
           IF "Z256_Manager".tOutputData.rgxDataToProcessInter[#TMP_dIndexFAST] THEN

               #TMP_dEncoderOverFAST_cmm := #TMP_dEncValueFast - "Z256_Manager".tOutputData.rgdFireHeadThreshold_cmm[#TMP_dIndexFAST];

               //firing
               IF #TMP_dEncoderOverFAST_cmm >= 0 THEN



                   IF ("Z256_Manager".tOutputData.rgxFireHeadON_OFF[#TMP_dIndexFAST]) AND ("M256_Manag_IDB".M256F_IDB[#TMP_dIndexFAST].ST_xOutputEnable) AND
                       "M256_Manag_IDB".M256M_ST_xAllHeadPositioned AND "M256_Manag_IDB".M256A_IDB[#TMP_dIndexFAST].OUTPUT_xCarriageDescent THEN

                       "M256_Manag_IDB".M256F_IDB[#TMP_dIndexFAST].OUTPUT_xFireON := 1;

                   ELSE

                       "M256_Manag_IDB".M256F_IDB[#TMP_dIndexFAST].OUTPUT_xFireON := 0;

                   END_IF;

                   #TMP_xChangeFAST := 1;
                   "Z256_Manager".tOutputData.rgxDataToProcessInter[#TMP_dIndexFAST] := 0;
                   "M256_Manag_IDB".M256F_IDB[#TMP_dIndexFAST].AUX_dHeadMissionIDinProg := "Z256_Manager".tOutputData.dMissionCode;
                   "M256_Manag_IDB".M256F_IDB[#TMP_dIndexFAST].AUX_xHeadFiringMissionInProgress := "Z256_Manager".tOutputData.rgxFireHeadON_OFF[#TMP_dIndexFAST];

                   #TMP_xDummy := false;
                   FOR #TMP_dIndexFAST_2 := 0 TO "CONST_dNumberOfHeadsCycle" DO
                       IF "Z256_Manager".tOutputData.rgxFireHeadON_OFF[#TMP_dIndexFAST_2] THEN
                           #TMP_xDummy := true;
                       END_IF;
                   END_FOR;
                   IF NOT (#TMP_xDummy) THEN
                       "M256_Manag_IDB".M256F_IDB[#TMP_dIndexFAST].AUX_dHeadMissionIDinProg := 0;
                   END_IF;
               END_IF;
           END_IF;
       END_FOR;


       #TMP_xDummy := false;
       FOR #TMP_dIndexFAST := 0 TO "CONST_dNumberOfHeadsCycle" DO
           IF "Z256_Manager".tOutputData.rgxDataToProcessInter[#TMP_dIndexFAST] <> 0 THEN
               #TMP_xDummy := true;
           END_IF;
       END_FOR;
       IF #TMP_xDummy = false THEN
           "Z256_Manager".tOutputData.xGateOpen := 0;
       END_IF;
       //Immagine di processo aggiornata automaticamente con l'OB
       //    IF #TMP_xChangeFAST THEN
       //        #TMP_iRetVal:=UPDAT_PO(PART := "IPP 1", FLADDR => "DEBUG_FiringAdressError");
       //    END_IF;


   END_IF;


   "o.1B160AP1.EnableCard1":=  "M256_Manag_IDB".M256F_IDB[0].OUTPUT_xFireON OR"M256_Manag_IDB".M256F_IDB[0].INPUT_xForceFiring;
   "o.1B160AP1.EnableCard2" := "M256_Manag_IDB".M256F_IDB[1].OUTPUT_xFireON OR "M256_Manag_IDB".M256F_IDB[1].INPUT_xForceFiring;
   "o.1B160AP1.EnableCard3" := "M256_Manag_IDB".M256F_IDB[2].OUTPUT_xFireON OR "M256_Manag_IDB".M256F_IDB[2].INPUT_xForceFiring;
   "o.1B160AP1.EnableCard4" := "M256_Manag_IDB".M256F_IDB[3].OUTPUT_xFireON OR "M256_Manag_IDB".M256F_IDB[3].INPUT_xForceFiring;
   "o.1B160AP1.EnableCard5" := "M256_Manag_IDB".M256F_IDB[4].OUTPUT_xFireON OR "M256_Manag_IDB".M256F_IDB[4].INPUT_xForceFiring;
   "o.1B160AP1.EnableCard5" := "M256_Manag_IDB".M256F_IDB[5].OUTPUT_xFireON OR "M256_Manag_IDB".M256F_IDB[4].INPUT_xForceFiring;
   "o.1B160AP1.EnableCard5" := "M256_Manag_IDB".M256F_IDB[6].OUTPUT_xFireON OR "M256_Manag_IDB".M256F_IDB[4].INPUT_xForceFiring;
   "o.1B160AP1.EnableCard5" := "M256_Manag_IDB".M256F_IDB[7].OUTPUT_xFireON OR "M256_Manag_IDB".M256F_IDB[4].INPUT_xForceFiring;
END_REGION
END_ORGANIZATION_BLOCK

ORGANIZATION_BLOCK "Startup"   // OB100, SCL, Startup
TITLE = "Complete Restart"
{ S7_Optimized_Access := 'TRUE' }
VERSION : 0.1
   VAR_INPUT
      LostRetentive : Bool;   // True if retentive data are lost
      LostRTC : Bool;   // True if date and time are lost
   END_VAR
   VAR_TEMP
      TMP_dIndex : DInt;
   END_VAR
BEGIN
   // Start Auto Sequence after PLC restart

   "OB_Initialize".IN_xInitialize := TRUE;

   "INIT_PlantCostants"();

   //FORCE MANUAL STATE
   "Z256_hmi".tHMW.xGeneralReset := 1;

   FOR #TMP_dIndex := 0 TO "CONST_dNumberOfHeadsCycle" DO
       "M256_Manag_IDB".M256M_IDB[#TMP_dIndex].ST_xHeadInitialized := 0;
       "M256_Manag_IDB".M256M_IDB[#TMP_dIndex].AUX_dHeadRequestPosition_cmm := "M256_Manag_IDB".M256M_IDB[#TMP_dIndex].tHMR.dHeadHomePositions_cmm; 
       "Z256_hmi".tHMW.rgxHeadEnabled[#TMP_dIndex] := true;
   END_FOR;
END_ORGANIZATION_BLOCK

// folder: 07_ArrayScada

FUNCTION "SCADA_Mapping" : Void   // FC8, SCL
{ S7_Optimized_Access := 'TRUE' }
VERSION : 0.1
   VAR_TEMP
      TMP_dIndex : DInt;
   END_VAR
BEGIN

   //Move Z256 HMR
   "DB_Z256_Scada".tHMR.xCalibrationsAllowed:="Z256_hmi".tHMR.xCalibrationsAllowed;
   "DB_Z256_Scada".tHMR.xZoneAlarm:="Z256_hmi".tHMR.xZoneAlarm;
   "DB_Z256_Scada".tHMR.dZoneMode:="Z256_hmi".tHMR.dZoneMode;

   "DB_Z256_Scada".tHMR.dCabinetStatusMCC:="Z256_hmi".tHMR.dCabinetStatus;
   "DB_Z256_Scada".tHMR.dProdModeRequest:="Z256_hmi".tHMR.dProdModeRequest;
   "DB_Z256_Scada".tHMR.dProdModeActual:="Z256_hmi".tHMR.dProdModeActual;

   "DB_Z256_Scada".tHMR."rgdHeadsActualStatus[0]":="Z256_hmi".tHMR.rgdHeadsActualStatus[0];
   "DB_Z256_Scada".tHMR."rgdHeadsActualStatus[1]":="Z256_hmi".tHMR.rgdHeadsActualStatus[1];
   "DB_Z256_Scada".tHMR."rgdHeadsActualStatus[2]":="Z256_hmi".tHMR.rgdHeadsActualStatus[2];
   "DB_Z256_Scada".tHMR."rgdHeadsActualStatus[3]":="Z256_hmi".tHMR.rgdHeadsActualStatus[3];
   "DB_Z256_Scada".tHMR."rgdHeadsActualStatus[4]":="Z256_hmi".tHMR.rgdHeadsActualStatus[4];
   "DB_Z256_Scada".tHMR."rgdHeadsActualStatus[5]":="Z256_hmi".tHMR.rgdHeadsActualStatus[5];
   "DB_Z256_Scada".tHMR."rgdHeadsActualStatus[6]":="Z256_hmi".tHMR.rgdHeadsActualStatus[6];
   "DB_Z256_Scada".tHMR."rgdHeadsActualStatus[7]":="Z256_hmi".tHMR.rgdHeadsActualStatus[7];


   //Move Z256 HMW
   //
   "Z256_hmi".tHMW.xFaultsReset:="DB_Z256_Scada".tHMW.xFaultsReset ;
   "Z256_hmi".tHMW.xAutoModeReq:= "DB_Z256_Scada".tHMW.xAutoModeReq ;
   "Z256_hmi".tHMW.xGeneralReset:= "DB_Z256_Scada".tHMW.xGeneralReset ;
   "Z256_hmi".tHMW.xCutOnBreakEnabled:="DB_Z256_Scada".tHMW.xCutOnBreakEnabled  ;
   "Z256_hmi".tHMW.xManModeReq := "DB_Z256_Scada".tHMW.xManModeReq;
   "Z256_hmi".tHMW.xMotorsAndCardsInitialize:= "DB_Z256_Scada".tHMW.xMotorsAndCardsInitialize ;
   "Z256_hmi".tHMW.xOutOfProdReq:= "DB_Z256_Scada".tHMW.xOutOfProdReq ;
   "Z256_hmi".tHMW.xInProdReq:= "DB_Z256_Scada".tHMW.xInProdReq   ;
   "Z256_hmi".tHMW.xPositionCalibrationRequest := "DB_Z256_Scada".tHMW.xPositionCalibrationRequest;
   "Z256_hmi".tHMW.xForceHeadsHoming:= "DB_Z256_Scada".tHMW.xForceHeadsHoming   ;
   "Z256_hmi".tHMW.xBridgeOffsetCalibrationRequest:="DB_Z256_Scada".tHMW.xBridgeOffsetCalibrationRequest;
   "Z256_hmi".tHMW.tManCmd.xBrakeEngage:="DB_Z256_Scada".tHMW.tManCmd.xBrakeEngage;
   "Z256_hmi".tHMW.tManCmd.xBrakeRelease:="DB_Z256_Scada".tHMW.tManCmd.xBrakeRelease;

   "Z256_hmi".tHMW.rgxHeadEnabled[0] := "DB_Z256_Scada".tHMW.xHeadEnabled_1;
   "Z256_hmi".tHMW.rgxHeadEnabled[1] := "DB_Z256_Scada".tHMW.xHeadEnabled_2;
   "Z256_hmi".tHMW.rgxHeadEnabled[2] := "DB_Z256_Scada".tHMW.xHeadEnabled_3;
   "Z256_hmi".tHMW.rgxHeadEnabled[3] := "DB_Z256_Scada".tHMW.xHeadEnabled_4;
   "Z256_hmi".tHMW.rgxHeadEnabled[4] := "DB_Z256_Scada".tHMW.xHeadEnabled_5;
   "Z256_hmi".tHMW.rgxHeadEnabled[5] := "DB_Z256_Scada".tHMW.xHeadEnabled_6;
   "Z256_hmi".tHMW.rgxHeadEnabled[6] := "DB_Z256_Scada".tHMW.xHeadEnabled_7;
   "Z256_hmi".tHMW.rgxHeadEnabled[7] := "DB_Z256_Scada".tHMW.xHeadEnabled_8;

   "Z256_hmi".tHMW.dMoveBridgeOffset_cmm := "DB_Z256_Scada".tHMW.dMoveBridgeOffset_cmm;
   "Z256_hmi".tHMW.dNumberOfLites := "DB_Z256_Scada".tHMW.dNumberOfLites;
   "Z256_hmi".tHMW.dPressureScalerOnSample_perc := "DB_Z256_Scada".tHMW.dPressureScalerOnSample_perc;

   "Z256_hmi".tHMW.rgdHeadSelected[0]:="DB_Z256_Scada".tHMW.dHead_Selected_1;
   "Z256_hmi".tHMW.rgdHeadSelected[1]:="DB_Z256_Scada".tHMW.dHead_Selected_2;
   "Z256_hmi".tHMW.rgdHeadSelected[2]:="DB_Z256_Scada".tHMW.dHead_Selected_3;
   "Z256_hmi".tHMW.rgdHeadSelected[3]:="DB_Z256_Scada".tHMW.dHead_Selected_4;
   "Z256_hmi".tHMW.rgdHeadSelected[4]:="DB_Z256_Scada".tHMW.dHead_Selected_5;
   "Z256_hmi".tHMW.rgdHeadSelected[5]:="DB_Z256_Scada".tHMW.dHead_Selected_6;
   "Z256_hmi".tHMW.rgdHeadSelected[6]:="DB_Z256_Scada".tHMW.dHead_Selected_7;
   "Z256_hmi".tHMW.rgdHeadSelected[7] :="DB_Z256_Scada".tHMW.dHead_Selected_8;

   "Z256_hmi".tHMW.rgdCutWidthTeo_cmm[0] := "DB_Z256_Scada".tHMW.dCutWidthTeo_cmm_1;
   "Z256_hmi".tHMW.rgdCutWidthTeo_cmm[1] := "DB_Z256_Scada".tHMW.dCutWidthTeo_cmm_2;
   "Z256_hmi".tHMW.rgdCutWidthTeo_cmm[2] := "DB_Z256_Scada".tHMW.dCutWidthTeo_cmm_3;
   "Z256_hmi".tHMW.rgdCutWidthTeo_cmm[3] := "DB_Z256_Scada".tHMW."dCutWidthTeo_cmm_4";
   "Z256_hmi".tHMW.rgdCutWidthTeo_cmm[4] := "DB_Z256_Scada".tHMW."dCutWidthTeo_cmm_5";
   "Z256_hmi".tHMW.rgdCutWidthTeo_cmm[5] := "DB_Z256_Scada".tHMW."dCutWidthTeo_cmm_6";
   "Z256_hmi".tHMW.rgdCutWidthTeo_cmm[6] := "DB_Z256_Scada".tHMW."dCutWidthTeo_cmm_7";
   "Z256_hmi".tHMW.rgdCutWidthTeo_cmm[7] := "DB_Z256_Scada".tHMW."dCutWidthTeo_cmm_8";


   "Z256_hmi".tHMW.rgdCutWidthReal_cmm[0]:="DB_Z256_Scada".tHMW.dCutWidthReal_cmm_1;
   "Z256_hmi".tHMW.rgdCutWidthReal_cmm[1]:="DB_Z256_Scada".tHMW.dCutWidthReal_cmm_2;
   "Z256_hmi".tHMW.rgdCutWidthReal_cmm[2]:="DB_Z256_Scada".tHMW.dCutWidthReal_cmm_3;
   "Z256_hmi".tHMW.rgdCutWidthReal_cmm[3]:="DB_Z256_Scada".tHMW."dCutWidthReal_cmm_4";
   "Z256_hmi".tHMW.rgdCutWidthReal_cmm[4]:="DB_Z256_Scada".tHMW."dCutWidthReal_cmm_5";
   "Z256_hmi".tHMW.rgdCutWidthReal_cmm[5]:="DB_Z256_Scada".tHMW."dCutWidthReal_cmm_6";
   "Z256_hmi".tHMW.rgdCutWidthReal_cmm[6]:="DB_Z256_Scada".tHMW."dCutWidthReal_cmm_7";
   "Z256_hmi".tHMW.rgdCutWidthReal_cmm[7]:="DB_Z256_Scada".tHMW."dCutWidthTeo_cmm_8";

   (* //Move Z256 ALM
   "DB_M256M_Scada".tAlm.tS.tS0 := "DB_Z256_Scada".tAlm.tS.tS0;
   "DB_Z256_Scada".tAlm.tS.tS0.x0 := "DB_Z256_Scada".tAlm.tS.tS0.x0;
   "DB_Z256_Scada".tAlm.tS.tS0.x1 := "DB_Z256_Scada".tAlm.tS.tS0.x1;
   "DB_Z256_Scada".tAlm.tS.tS0.x2 := "DB_Z256_Scada".tAlm.tS.tS0.x2;
   "DB_Z256_Scada".tAlm.tS.tS0.x3 := "DB_Z256_Scada".tAlm.tS.tS0.x3;
   "DB_Z256_Scada".tAlm.tS.tS0.x4 := "DB_Z256_Scada".tAlm.tS.tS0.x4;
   "DB_Z256_Scada".tAlm.tS.tS0.x5 := "DB_Z256_Scada".tAlm.tS.tS0.x5;
   "DB_Z256_Scada".tAlm.tS.tS0.x6 := "DB_Z256_Scada".tAlm.tS.tS0.x6;
   "DB_Z256_Scada".tAlm.tS.tS0.x7 := "DB_Z256_Scada".tAlm.tS.tS0.x7;
   "DB_Z256_Scada".tAlm.tS.tS0.x8 := "DB_Z256_Scada".tAlm.tS.tS0.x8;

   "DB_Z256_Scada".tAlm.tS.tS0.x9 := "DB_Z256_Scada".tAlm.tS.tS0.x9;
   "DB_Z256_Scada".tAlm.tS.tS0.x10 := "DB_Z256_Scada".tAlm.tS.tS0.x10;
   "DB_Z256_Scada".tAlm.tS.tS0.x11 := "DB_Z256_Scada".tAlm.tS.tS0.x11;
   "DB_Z256_Scada".tAlm.tS.tS0.x12 := "DB_Z256_Scada".tAlm.tS.tS0.x12;
   "DB_Z256_Scada".tAlm.tS.tS0.x13 := "DB_Z256_Scada".tAlm.tS.tS0.x13;
   "DB_Z256_Scada".tAlm.tS.tS0.x14 := "DB_Z256_Scada".tAlm.tS.tS0.x14;
   "DB_Z256_Scada".tAlm.tS.tS0.x15 := "DB_Z256_Scada".tAlm.tS.tS0.x15;
   "DB_Z256_Scada".tAlm.tS.tS0.x16 := "DB_Z256_Scada".tAlm.tS.tS0.x16;
   "DB_Z256_Scada".tAlm.tS.tS0.x17 := "DB_Z256_Scada".tAlm.tS.tS0.x17;

   "DB_Z256_Scada".tAlm.tS.tS0.x18 := "DB_Z256_Scada".tAlm.tS.tS0.x18;
   "DB_Z256_Scada".tAlm.tS.tS0.x19 := "DB_Z256_Scada".tAlm.tS.tS0.x19;
   "DB_Z256_Scada".tAlm.tS.tS0.x20 := "DB_Z256_Scada".tAlm.tS.tS0.x20;
   "DB_Z256_Scada".tAlm.tS.tS0.x21 := "DB_Z256_Scada".tAlm.tS.tS0.x21;
   "DB_Z256_Scada".tAlm.tS.tS0.x22 := "DB_Z256_Scada".tAlm.tS.tS0.x22;
   "DB_Z256_Scada".tAlm.tS.tS0.x23 := "DB_Z256_Scada".tAlm.tS.tS0.x23;
   "DB_Z256_Scada".tAlm.tS.tS0.x24 := "DB_Z256_Scada".tAlm.tS.tS0.x24;
   "DB_Z256_Scada".tAlm.tS.tS0.x25 := "DB_Z256_Scada".tAlm.tS.tS0.x25;
   "DB_Z256_Scada".tAlm.tS.tS0.x26 := "DB_Z256_Scada".tAlm.tS.tS0.x26;
   "DB_Z256_Scada".tAlm.tS.tS0.x27 := "DB_Z256_Scada".tAlm.tS.tS0.x27;
   "DB_Z256_Scada".tAlm.tS.tS0.x28 := "DB_Z256_Scada".tAlm.tS.tS0.x28;
   "DB_Z256_Scada".tAlm.tS.tS0.x29 := "DB_Z256_Scada".tAlm.tS.tS0.x29;
   "DB_Z256_Scada".tAlm.tS.tS0.x30 := "DB_Z256_Scada".tAlm.tS.tS0.x30;
   "DB_Z256_Scada".tAlm.tS.tS0.x31 := "DB_Z256_Scada".tAlm.tS.tS0.x31; *)


    //Move M256M MOVEMENTS HMR
    //H1
   "DB_M256M_Scada".tHMR.tManCmd.xManJogForwardFdbk_H1 := "M256_Manag_IDB".M256M_IDB[0].tHMR.tManCmd.xMan_JogForwardFdbk;
   "DB_M256M_Scada".tHMR.tManCmd.xManJogBackwardFdbk_H1 := "M256_Manag_IDB".M256M_IDB[0].tHMR.tManCmd.xMan_JogBackwardFdbk;
   "DB_M256M_Scada".tHMR.iCodeAlarm_H1 := "M256_Manag_IDB".M256M_IDB[0].tHMR.iCodeAlarm;
   "DB_M256M_Scada".tHMR.dHeadActualPositions_cmm_H1 := "M256_Manag_IDB".M256M_IDB[0].tHMR.dHeadActualPositions_cmm;
   "DB_M256M_Scada".tHMR.dHeadHomePositions_cmm_H1 := "M256_Manag_IDB".M256M_IDB[0].tHMR.dHeadHomePositions_cmm;
   "DB_M256M_Scada".tHMR.dHeadMoveStatus_H1 := "M256_Manag_IDB".M256M_IDB[0].tHMR.rgdHeadMoveStatus;
   //H2 
   "DB_M256M_Scada".tHMR.tManCmd.xManJogBackwardFdbk_H2 := "M256_Manag_IDB".M256M_IDB[1].tHMR.tManCmd.xMan_JogForwardFdbk;
   "DB_M256M_Scada".tHMR.tManCmd.xManJogBackwardFdbk_H2 := "M256_Manag_IDB".M256M_IDB[1].tHMR.tManCmd.xMan_JogBackwardFdbk;
   "DB_M256M_Scada".tHMR.iCodeAlarm_H2 := "M256_Manag_IDB".M256M_IDB[1].tHMR.iCodeAlarm;
   "DB_M256M_Scada".tHMR.dHeadActualPositions_cmm_H2 := "M256_Manag_IDB".M256M_IDB[1].tHMR.dHeadActualPositions_cmm;
   "DB_M256M_Scada".tHMR.dHeadHomePositions_cmm_H2 := "M256_Manag_IDB".M256M_IDB[1].tHMR.dHeadHomePositions_cmm;
   "DB_M256M_Scada".tHMR.dHeadMoveStatus_H2 := "M256_Manag_IDB".M256M_IDB[1].tHMR.rgdHeadMoveStatus;
   //H3 
   "DB_M256M_Scada".tHMR.tManCmd.xManJogForwardFdbk_H3 :="M256_Manag_IDB".M256M_IDB[2].tHMR.tManCmd.xMan_JogForwardFdbk;
   "DB_M256M_Scada".tHMR.tManCmd.xManJogBackwardFdbk_H3 := "M256_Manag_IDB".M256M_IDB[2].tHMR.tManCmd.xMan_JogBackwardFdbk;
   "DB_M256M_Scada".tHMR.iCodeAlarm_H3 := "M256_Manag_IDB".M256M_IDB[2].tHMR.iCodeAlarm;
   "DB_M256M_Scada".tHMR.dHeadActualPositions_cmm_H3 := "M256_Manag_IDB".M256M_IDB[2].tHMR.dHeadActualPositions_cmm;
   "DB_M256M_Scada".tHMR.dHeadHomePositions_cmm_H3 := "M256_Manag_IDB".M256M_IDB[2].tHMR.dHeadHomePositions_cmm;
   "DB_M256M_Scada".tHMR.dHeadMoveStatus_H3 := "M256_Manag_IDB".M256M_IDB[2].tHMR.rgdHeadMoveStatus;
   //H4 
   "DB_M256M_Scada".tHMR.tManCmd.xManJogForwardFdbk_H4:= "M256_Manag_IDB".M256M_IDB[3].tHMR.tManCmd.xMan_JogForwardFdbk;
   "DB_M256M_Scada".tHMR.tManCmd.xManJogBackwardFdbk_H4 := "M256_Manag_IDB".M256M_IDB[3].tHMR.tManCmd.xMan_JogBackwardFdbk;
   "DB_M256M_Scada".tHMR.iCodeAlarm_H4 := "M256_Manag_IDB".M256M_IDB[3].tHMR.iCodeAlarm;
   "DB_M256M_Scada".tHMR.dHeadActualPositions_cmm_H4 := "M256_Manag_IDB".M256M_IDB[3].tHMR.dHeadActualPositions_cmm;
   "DB_M256M_Scada".tHMR.dHeadHomePositions_cmm_H4 := "M256_Manag_IDB".M256M_IDB[3].tHMR.dHeadHomePositions_cmm;
   "DB_M256M_Scada".tHMR.dHeadMoveStatus_H4 := "M256_Manag_IDB".M256M_IDB[3].tHMR.rgdHeadMoveStatus;
   "DB_M256M_Scada".tHMR.iCodeAlarm_H4 := "M256_Manag_IDB".M256M_IDB[3].tHMR.iCodeAlarm;
   //H5
   "DB_M256M_Scada".tHMR.tManCmd.xManJogForwardFdbk_H5 := "M256_Manag_IDB".M256M_IDB[4].tHMR.tManCmd.xMan_JogForwardFdbk;
   "DB_M256M_Scada".tHMR.tManCmd.xManJogBackwardFdbk_H5:= "M256_Manag_IDB".M256M_IDB[4].tHMR.tManCmd.xMan_JogBackwardFdbk;
   "DB_M256M_Scada".tHMR.iCodeAlarm_H5 := "M256_Manag_IDB".M256M_IDB[4].tHMR.iCodeAlarm;
   "DB_M256M_Scada".tHMR.dHeadActualPositions_cmm_H5 := "M256_Manag_IDB".M256M_IDB[4].tHMR.dHeadActualPositions_cmm;
   "DB_M256M_Scada".tHMR.dHeadHomePositions_cmm_H5 := "M256_Manag_IDB".M256M_IDB[4].tHMR.dHeadHomePositions_cmm;
   "DB_M256M_Scada".tHMR.dHeadMoveStatus_H5 := "M256_Manag_IDB".M256M_IDB[4].tHMR.rgdHeadMoveStatus;
   //H6 
   "DB_M256M_Scada".tHMR.tManCmd.xManJogForwardFdbk_H6 := "M256_Manag_IDB".M256M_IDB[5].tHMR.tManCmd.xMan_JogForwardFdbk;
   "DB_M256M_Scada".tHMR.tManCmd.xManJogBackwardFdbk_H6 := "M256_Manag_IDB".M256M_IDB[5].tHMR.tManCmd.xMan_JogBackwardFdbk;
   "DB_M256M_Scada".tHMR.iCodeAlarm_H6 := "M256_Manag_IDB".M256M_IDB[5].tHMR.iCodeAlarm;
   "DB_M256M_Scada".tHMR.dHeadActualPositions_cmm_H6 := "M256_Manag_IDB".M256M_IDB[5].tHMR.dHeadActualPositions_cmm;
   "DB_M256M_Scada".tHMR.dHeadHomePositions_cmm_H6 := "M256_Manag_IDB".M256M_IDB[5].tHMR.dHeadHomePositions_cmm;
   "DB_M256M_Scada".tHMR.dHeadMoveStatus_H6 := "M256_Manag_IDB".M256M_IDB[5].tHMR.rgdHeadMoveStatus;
   //H7 
   "DB_M256M_Scada".tHMR.tManCmd.xManJogForwardFdbk_H7 := "M256_Manag_IDB".M256M_IDB[6].tHMR.tManCmd.xMan_JogForwardFdbk;
   "DB_M256M_Scada".tHMR.tManCmd.xManJogBackwardFdbk_H7 := "M256_Manag_IDB".M256M_IDB[6].tHMR.tManCmd.xMan_JogBackwardFdbk;
   "DB_M256M_Scada".tHMR.iCodeAlarm_H7 := "M256_Manag_IDB".M256M_IDB[6].tHMR.iCodeAlarm;
   "DB_M256M_Scada".tHMR.dHeadActualPositions_cmm_H7 := "M256_Manag_IDB".M256M_IDB[6].tHMR.dHeadActualPositions_cmm;
   "DB_M256M_Scada".tHMR.dHeadHomePositions_cmm_H7 := "M256_Manag_IDB".M256M_IDB[6].tHMR.dHeadHomePositions_cmm;
   "DB_M256M_Scada".tHMR.dHeadMoveStatus_H7 := "M256_Manag_IDB".M256M_IDB[6].tHMR.rgdHeadMoveStatus;
   //H8 
   "DB_M256M_Scada".tHMR.tManCmd.xManJogForwardFdbk_H8 := "M256_Manag_IDB".M256M_IDB[7].tHMR.tManCmd.xMan_JogForwardFdbk;
   "DB_M256M_Scada".tHMR.tManCmd.xManJogBackwardFdbk_H8 := "M256_Manag_IDB".M256M_IDB[7].tHMR.tManCmd.xMan_JogBackwardFdbk;
   "DB_M256M_Scada".tHMR.iCodeAlarm_H8 := "M256_Manag_IDB".M256M_IDB[7].tHMR.iCodeAlarm;
   "DB_M256M_Scada".tHMR.dHeadActualPositions_cmm_H8 := "M256_Manag_IDB".M256M_IDB[7].tHMR.dHeadActualPositions_cmm;
   "DB_M256M_Scada".tHMR.dHeadHomePositions_cmm_H8 := "M256_Manag_IDB".M256M_IDB[7].tHMR.dHeadHomePositions_cmm;
   "DB_M256M_Scada".tHMR.dHeadMoveStatus_H8 := "M256_Manag_IDB".M256M_IDB[7].tHMR.rgdHeadMoveStatus;


       //Move MOVEMENTS HMW

       //H1
       "M256_Manag_IDB".M256M_IDB[0].tHMW.dHeadHomePositions_cmm := "DB_M256M_Scada".tHMW.dHeadHomePositions_cmm_H1;
       "M256_Manag_IDB".M256M_IDB[0].tHMW.xBrakeEngageHeads := "DB_M256M_Scada".tHMW.xBrakeRealeaseHead_H1;
       "M256_Manag_IDB".M256M_IDB[0].tHMW.xBrakeRealeaseHeads := "DB_M256M_Scada".tHMW.xBrakeEngageHeads_H1;
       "M256_Manag_IDB".M256M_IDB[0].tHMW.xUpdateHomeHead := "DB_M256M_Scada".tHMW.xUpdateHomeHead_H1;
       "M256_Manag_IDB".M256M_IDB[0].tHMW.tManCmd.xMan_JogBackward := "DB_M256M_Scada".tHMW.tManCmd.xMan_JogBackward_H1;
       "M256_Manag_IDB".M256M_IDB[0].tHMW.tManCmd.xMan_JogForward := "DB_M256M_Scada".tHMW.tManCmd.xMan_JogForward_H1;
       //H2
       "M256_Manag_IDB".M256M_IDB[1].tHMW.dHeadHomePositions_cmm := "DB_M256M_Scada".tHMW.dHeadHomePositions_cmm_H2;
       "M256_Manag_IDB".M256M_IDB[1].tHMW.xBrakeEngageHeads := "DB_M256M_Scada".tHMW.xBrakeRealeaseHead_H2;
       "M256_Manag_IDB".M256M_IDB[1].tHMW.xBrakeRealeaseHeads := "DB_M256M_Scada".tHMW.xBrakeEngageHeads_H2;
       "M256_Manag_IDB".M256M_IDB[1].tHMW.xUpdateHomeHead := "DB_M256M_Scada".tHMW.xUpdateHomeHead_H2;
       "M256_Manag_IDB".M256M_IDB[1].tHMW.tManCmd.xMan_JogBackward := "DB_M256M_Scada".tHMW.tManCmd.xMan_JogBackward_H2;
       "M256_Manag_IDB".M256M_IDB[1].tHMW.tManCmd.xMan_JogForward := "DB_M256M_Scada".tHMW.tManCmd.xMan_JogForward_H2;
       //H3
       "M256_Manag_IDB".M256M_IDB[2].tHMW.dHeadHomePositions_cmm := "DB_M256M_Scada".tHMW.dHeadHomePositions_cmm_H3;
       "M256_Manag_IDB".M256M_IDB[2].tHMW.xBrakeEngageHeads := "DB_M256M_Scada".tHMW.xBrakeRealeaseHead_H3;
       "M256_Manag_IDB".M256M_IDB[2].tHMW.xBrakeRealeaseHeads := "DB_M256M_Scada".tHMW.xBrakeEngageHeads_H3;
       "M256_Manag_IDB".M256M_IDB[2].tHMW.xUpdateHomeHead := "DB_M256M_Scada".tHMW.xUpdateHomeHead_H3;
       "M256_Manag_IDB".M256M_IDB[2].tHMW.tManCmd.xMan_JogBackward := "DB_M256M_Scada".tHMW.tManCmd.xMan_JogBackward_H3;
       "M256_Manag_IDB".M256M_IDB[2].tHMW.tManCmd.xMan_JogForward := "DB_M256M_Scada".tHMW.tManCmd.xMan_JogForward_H3;
       //H4
       "M256_Manag_IDB".M256M_IDB[3].tHMW.dHeadHomePositions_cmm := "DB_M256M_Scada".tHMW.dHeadHomePositions_cmm_H4;
       "M256_Manag_IDB".M256M_IDB[3].tHMW.xBrakeEngageHeads := "DB_M256M_Scada".tHMW.xBrakeRealeaseHead_H4;
       "M256_Manag_IDB".M256M_IDB[3].tHMW.xBrakeRealeaseHeads := "DB_M256M_Scada".tHMW.xBrakeEngageHeads_H4;
       "M256_Manag_IDB".M256M_IDB[3].tHMW.xUpdateHomeHead := "DB_M256M_Scada".tHMW.xUpdateHomeHead_H4;
       "M256_Manag_IDB".M256M_IDB[3].tHMW.tManCmd.xMan_JogBackward := "DB_M256M_Scada".tHMW.tManCmd.xMan_JogBackward_H4;
       "M256_Manag_IDB".M256M_IDB[3].tHMW.tManCmd.xMan_JogForward := "DB_M256M_Scada".tHMW.tManCmd.xMan_JogForward_H4;
       //H5
       "M256_Manag_IDB".M256M_IDB[4].tHMW.dHeadHomePositions_cmm := "DB_M256M_Scada".tHMW.dHeadHomePositions_cmm_H5;
       "M256_Manag_IDB".M256M_IDB[4].tHMW.xBrakeEngageHeads := "DB_M256M_Scada".tHMW.xBrakeRealeaseHead_H5;
       "M256_Manag_IDB".M256M_IDB[4].tHMW.xBrakeRealeaseHeads := "DB_M256M_Scada".tHMW.xBrakeEngageHeads_H5;
       "M256_Manag_IDB".M256M_IDB[4].tHMW.xUpdateHomeHead := "DB_M256M_Scada".tHMW.xUpdateHomeHead_H5;
       "M256_Manag_IDB".M256M_IDB[4].tHMW.tManCmd.xMan_JogBackward := "DB_M256M_Scada".tHMW.tManCmd.xMan_JogBackward_H5;
       "M256_Manag_IDB".M256M_IDB[4].tHMW.tManCmd.xMan_JogForward := "DB_M256M_Scada".tHMW.tManCmd.xMan_JogForward_H5;
       //H6
       "M256_Manag_IDB".M256M_IDB[5].tHMW.dHeadHomePositions_cmm := "DB_M256M_Scada".tHMW.dHeadHomePositions_cmm_H6;
       "M256_Manag_IDB".M256M_IDB[5].tHMW.xBrakeEngageHeads := "DB_M256M_Scada".tHMW.xBrakeRealeaseHead_H6;
       "M256_Manag_IDB".M256M_IDB[5].tHMW.xBrakeRealeaseHeads := "DB_M256M_Scada".tHMW.xBrakeEngageHeads_H6;
       "M256_Manag_IDB".M256M_IDB[5].tHMW.xUpdateHomeHead := "DB_M256M_Scada".tHMW.xUpdateHomeHead_H6;
       "M256_Manag_IDB".M256M_IDB[5].tHMW.tManCmd.xMan_JogBackward := "DB_M256M_Scada".tHMW.tManCmd.xMan_JogBackward_H6;
       "M256_Manag_IDB".M256M_IDB[5].tHMW.tManCmd.xMan_JogForward := "DB_M256M_Scada".tHMW.tManCmd.xMan_JogForward_H6;
       //H7
       "M256_Manag_IDB".M256M_IDB[6].tHMW.dHeadHomePositions_cmm := "DB_M256M_Scada".tHMW.dHeadHomePositions_cmm_H7;
       "M256_Manag_IDB".M256M_IDB[6].tHMW.xBrakeEngageHeads := "DB_M256M_Scada".tHMW.xBrakeRealeaseHead_H7;
       "M256_Manag_IDB".M256M_IDB[6].tHMW.xBrakeRealeaseHeads := "DB_M256M_Scada".tHMW.xBrakeEngageHeads_H7;
       "M256_Manag_IDB".M256M_IDB[6].tHMW.xUpdateHomeHead := "DB_M256M_Scada".tHMW.xUpdateHomeHead_H7;
       "M256_Manag_IDB".M256M_IDB[6].tHMW.tManCmd.xMan_JogBackward := "DB_M256M_Scada".tHMW.tManCmd.xMan_JogBackward_H7;
       "M256_Manag_IDB".M256M_IDB[6].tHMW.tManCmd.xMan_JogForward := "DB_M256M_Scada".tHMW.tManCmd.xMan_JogForward_H7;

       //H8
       "M256_Manag_IDB".M256M_IDB[7].tHMW.dHeadHomePositions_cmm := "DB_M256M_Scada".tHMW.dHeadHomePositions_cmm_H8;
       "M256_Manag_IDB".M256M_IDB[7].tHMW.xBrakeEngageHeads := "DB_M256M_Scada".tHMW.xBrakeRealeaseHead_H8;
       "M256_Manag_IDB".M256M_IDB[7].tHMW.xBrakeRealeaseHeads := "DB_M256M_Scada".tHMW.xBrakeEngageHeads_H8;
       "M256_Manag_IDB".M256M_IDB[7].tHMW.xUpdateHomeHead := "DB_M256M_Scada".tHMW.xUpdateHomeHead_H8;
       "M256_Manag_IDB".M256M_IDB[7].tHMW.tManCmd.xMan_JogBackward := "DB_M256M_Scada".tHMW.tManCmd.xMan_JogBackward_H8;
       "M256_Manag_IDB".M256M_IDB[7].tHMW.tManCmd.xMan_JogForward := "DB_M256M_Scada".tHMW.tManCmd.xMan_JogForward_H8;

       //Move MOVEMENTS ALM
       //H1
       "DB_M256M_Scada".tAlm.tS.tS0.x0 := "M256_Manag_IDB".M256M_IDB[0].tALM.tS.x0;
       "DB_M256M_Scada".tAlm.tS.tS0.x1 := "M256_Manag_IDB".M256M_IDB[0].tALM.tS.x1;
       "DB_M256M_Scada".tAlm.tS.tS0.x2 := "M256_Manag_IDB".M256M_IDB[0].tALM.tS.x2;
       "DB_M256M_Scada".tAlm.tS.tS0.x3 := "M256_Manag_IDB".M256M_IDB[0].tALM.tS.x3;
       "DB_M256M_Scada".tAlm.tS.tS0.x4 := "M256_Manag_IDB".M256M_IDB[0].tALM.tS.x4;
       "DB_M256M_Scada".tAlm.tS.tS0.x5 := "M256_Manag_IDB".M256M_IDB[0].tALM.tS.x5;
       "DB_M256M_Scada".tAlm.tS.tS0.x6 := "M256_Manag_IDB".M256M_IDB[0].tALM.tS.x6;
       "DB_M256M_Scada".tAlm.tS.tS0.x7 := "M256_Manag_IDB".M256M_IDB[0].tALM.tS.x7;
       "DB_M256M_Scada".tAlm.tS.tS0.x8 := "M256_Manag_IDB".M256M_IDB[0].tALM.tS.x8;
       //H2
       "DB_M256M_Scada".tAlm.tS.tS0.x9 := "M256_Manag_IDB".M256M_IDB[1].tALM.tS.x0;
       "DB_M256M_Scada".tAlm.tS.tS0.x10 := "M256_Manag_IDB".M256M_IDB[1].tALM.tS.x1;
       "DB_M256M_Scada".tAlm.tS.tS0.x11 := "M256_Manag_IDB".M256M_IDB[1].tALM.tS.x2;
       "DB_M256M_Scada".tAlm.tS.tS0.x12 := "M256_Manag_IDB".M256M_IDB[1].tALM.tS.x3;
       "DB_M256M_Scada".tAlm.tS.tS0.x13 := "M256_Manag_IDB".M256M_IDB[1].tALM.tS.x4;
       "DB_M256M_Scada".tAlm.tS.tS0.x14 := "M256_Manag_IDB".M256M_IDB[1].tALM.tS.x5;
       "DB_M256M_Scada".tAlm.tS.tS0.x15 := "M256_Manag_IDB".M256M_IDB[1].tALM.tS.x6;
       "DB_M256M_Scada".tAlm.tS.tS0.x16 := "M256_Manag_IDB".M256M_IDB[1].tALM.tS.x7;
       "DB_M256M_Scada".tAlm.tS.tS0.x17 := "M256_Manag_IDB".M256M_IDB[1].tALM.tS.x8;
       //H3
       "DB_M256M_Scada".tAlm.tS.tS0.x18 := "M256_Manag_IDB".M256M_IDB[2].tALM.tS.x0;
       "DB_M256M_Scada".tAlm.tS.tS0.x19 := "M256_Manag_IDB".M256M_IDB[2].tALM.tS.x1;
       "DB_M256M_Scada".tAlm.tS.tS0.x20 := "M256_Manag_IDB".M256M_IDB[2].tALM.tS.x2;
       "DB_M256M_Scada".tAlm.tS.tS0.x21 := "M256_Manag_IDB".M256M_IDB[2].tALM.tS.x3;
       "DB_M256M_Scada".tAlm.tS.tS0.x22 := "M256_Manag_IDB".M256M_IDB[2].tALM.tS.x4;
       "DB_M256M_Scada".tAlm.tS.tS0.x23 := "M256_Manag_IDB".M256M_IDB[2].tALM.tS.x5;
       "DB_M256M_Scada".tAlm.tS.tS0.x24 := "M256_Manag_IDB".M256M_IDB[2].tALM.tS.x6;
       "DB_M256M_Scada".tAlm.tS.tS0.x25 := "M256_Manag_IDB".M256M_IDB[2].tALM.tS.x7;
       "DB_M256M_Scada".tAlm.tS.tS0.x26 := "M256_Manag_IDB".M256M_IDB[2].tALM.tS.x8;
       //H4
       "DB_M256M_Scada".tAlm.tS.tS1.x0 := "M256_Manag_IDB".M256M_IDB[3].tALM.tS.x0;
       "DB_M256M_Scada".tAlm.tS.tS1.x1 := "M256_Manag_IDB".M256M_IDB[3].tALM.tS.x1;
       "DB_M256M_Scada".tAlm.tS.tS1.x2 := "M256_Manag_IDB".M256M_IDB[3].tALM.tS.x2;
       "DB_M256M_Scada".tAlm.tS.tS1.x3 := "M256_Manag_IDB".M256M_IDB[3].tALM.tS.x3;
       "DB_M256M_Scada".tAlm.tS.tS1.x4 := "M256_Manag_IDB".M256M_IDB[3].tALM.tS.x4;
       "DB_M256M_Scada".tAlm.tS.tS1.x5 := "M256_Manag_IDB".M256M_IDB[3].tALM.tS.x5;
       "DB_M256M_Scada".tAlm.tS.tS1.x6 := "M256_Manag_IDB".M256M_IDB[3].tALM.tS.x6;
       "DB_M256M_Scada".tAlm.tS.tS1.x7 := "M256_Manag_IDB".M256M_IDB[3].tALM.tS.x7;
       "DB_M256M_Scada".tAlm.tS.tS1.x8 := "M256_Manag_IDB".M256M_IDB[3].tALM.tS.x8;
       //H5
       "DB_M256M_Scada".tAlm.tS.tS1.x9 := "M256_Manag_IDB".M256M_IDB[4].tALM.tS.x0;
       "DB_M256M_Scada".tAlm.tS.tS1.x10 := "M256_Manag_IDB".M256M_IDB[4].tALM.tS.x1;
       "DB_M256M_Scada".tAlm.tS.tS1.x11 := "M256_Manag_IDB".M256M_IDB[4].tALM.tS.x2;
       "DB_M256M_Scada".tAlm.tS.tS1.x12 := "M256_Manag_IDB".M256M_IDB[4].tALM.tS.x3;
       "DB_M256M_Scada".tAlm.tS.tS1.x13 := "M256_Manag_IDB".M256M_IDB[4].tALM.tS.x4;
       "DB_M256M_Scada".tAlm.tS.tS1.x14 := "M256_Manag_IDB".M256M_IDB[4].tALM.tS.x5;
       "DB_M256M_Scada".tAlm.tS.tS1.x15 := "M256_Manag_IDB".M256M_IDB[4].tALM.tS.x6;
       "DB_M256M_Scada".tAlm.tS.tS1.x16 := "M256_Manag_IDB".M256M_IDB[4].tALM.tS.x7;
       "DB_M256M_Scada".tAlm.tS.tS1.x17 := "M256_Manag_IDB".M256M_IDB[4].tALM.tS.x8;
       //H6
       "DB_M256M_Scada".tAlm.tS.tS1.x18 := "M256_Manag_IDB".M256M_IDB[5].tALM.tS.x0;
       "DB_M256M_Scada".tAlm.tS.tS1.x19 := "M256_Manag_IDB".M256M_IDB[5].tALM.tS.x1;
       "DB_M256M_Scada".tAlm.tS.tS1.x20 := "M256_Manag_IDB".M256M_IDB[5].tALM.tS.x2;
       "DB_M256M_Scada".tAlm.tS.tS1.x21 := "M256_Manag_IDB".M256M_IDB[5].tALM.tS.x3;
       "DB_M256M_Scada".tAlm.tS.tS1.x22 := "M256_Manag_IDB".M256M_IDB[5].tALM.tS.x4;
       "DB_M256M_Scada".tAlm.tS.tS1.x23 := "M256_Manag_IDB".M256M_IDB[5].tALM.tS.x5;
       "DB_M256M_Scada".tAlm.tS.tS1.x24 := "M256_Manag_IDB".M256M_IDB[5].tALM.tS.x6;
       "DB_M256M_Scada".tAlm.tS.tS1.x25 := "M256_Manag_IDB".M256M_IDB[5].tALM.tS.x7;
       "DB_M256M_Scada".tAlm.tS.tS1.x26 := "M256_Manag_IDB".M256M_IDB[5].tALM.tS.x8;
       //H7
       "DB_M256M_Scada".tAlm.tS.tS2.x0 := "M256_Manag_IDB".M256M_IDB[6].tALM.tS.x0;
       "DB_M256M_Scada".tAlm.tS.tS2.x1 := "M256_Manag_IDB".M256M_IDB[6].tALM.tS.x1;
       "DB_M256M_Scada".tAlm.tS.tS2.x2 := "M256_Manag_IDB".M256M_IDB[6].tALM.tS.x2;
       "DB_M256M_Scada".tAlm.tS.tS2.x3 := "M256_Manag_IDB".M256M_IDB[6].tALM.tS.x3;
       "DB_M256M_Scada".tAlm.tS.tS2.x4 := "M256_Manag_IDB".M256M_IDB[6].tALM.tS.x4;
       "DB_M256M_Scada".tAlm.tS.tS2.x5 := "M256_Manag_IDB".M256M_IDB[6].tALM.tS.x5;
       "DB_M256M_Scada".tAlm.tS.tS2.x6 := "M256_Manag_IDB".M256M_IDB[6].tALM.tS.x6;
       "DB_M256M_Scada".tAlm.tS.tS2.x7 := "M256_Manag_IDB".M256M_IDB[6].tALM.tS.x7;
       "DB_M256M_Scada".tAlm.tS.tS2.x8 := "M256_Manag_IDB".M256M_IDB[6].tALM.tS.x8;
       //H8
       "DB_M256M_Scada".tAlm.tS.tS2.x9 := "M256_Manag_IDB".M256M_IDB[7].tALM.tS.x0;
       "DB_M256M_Scada".tAlm.tS.tS2.x10 := "M256_Manag_IDB".M256M_IDB[7].tALM.tS.x1;
       "DB_M256M_Scada".tAlm.tS.tS2.x11 := "M256_Manag_IDB".M256M_IDB[7].tALM.tS.x2;
       "DB_M256M_Scada".tAlm.tS.tS2.x12:= "M256_Manag_IDB".M256M_IDB[7].tALM.tS.x3;
       "DB_M256M_Scada".tAlm.tS.tS2.x13 := "M256_Manag_IDB".M256M_IDB[7].tALM.tS.x4;
       "DB_M256M_Scada".tAlm.tS.tS2.x14 := "M256_Manag_IDB".M256M_IDB[7].tALM.tS.x5;
       "DB_M256M_Scada".tAlm.tS.tS2.x15 := "M256_Manag_IDB".M256M_IDB[7].tALM.tS.x6;
       "DB_M256M_Scada".tAlm.tS.tS2.x16 := "M256_Manag_IDB".M256M_IDB[7].tALM.tS.x7;
       "DB_M256M_Scada".tAlm.tS.tS2.x17 := "M256_Manag_IDB".M256M_IDB[7].tALM.tS.x8;


       //Move FIRE HMR
       //H1
       "DB_M256F_Scada".tHMR.dHeadStatus_H1 := "M256_Manag_IDB".M256F_IDB[0].tHMR.dHeadStatus;
       "DB_M256F_Scada".tHMR.rHeadUsage_km_H1 := "M256_Manag_IDB".M256F_IDB[0].tHMR.rHeadUsage_km;
       "DB_M256F_Scada".tHMR.tManCmd.xMan_FireON_Fdbk_H1 := "M256_Manag_IDB".M256F_IDB[0].tHMR.tManCmd.xMan_FireON_Fdbk;
       "DB_M256F_Scada".tHMR.tManCmd.xMan_FireOFF_Fdbk_H1 := "M256_Manag_IDB".M256F_IDB[0].tHMR.tManCmd.xMan_FireOFF_Fdbk;
       "DB_M256F_Scada".tHMR.tManCmd.xMan_OilON_Fdbk_H1 := "M256_Manag_IDB".M256F_IDB[0].tHMR.tManCmd.xMan_OilON_Fdbk;

       //H2
       "DB_M256F_Scada".tHMR.dHeadStatus_H2 := "M256_Manag_IDB".M256F_IDB[1].tHMR.dHeadStatus;
       "DB_M256F_Scada".tHMR.rHeadUsage_km_H2 := "M256_Manag_IDB".M256F_IDB[1].tHMR.rHeadUsage_km;
       "DB_M256F_Scada".tHMR.tManCmd.xMan_FireON_Fdbk_H2 := "M256_Manag_IDB".M256F_IDB[1].tHMR.tManCmd.xMan_FireON_Fdbk;
       "DB_M256F_Scada".tHMR.tManCmd.xMan_FireOFF_Fdbk_H2 := "M256_Manag_IDB".M256F_IDB[1].tHMR.tManCmd.xMan_FireOFF_Fdbk;
       "DB_M256F_Scada".tHMR.tManCmd.xMan_OilON_Fdbk_H2 := "M256_Manag_IDB".M256F_IDB[1].tHMR.tManCmd.xMan_OilON_Fdbk;

       //H3
       "DB_M256F_Scada".tHMR.dHeadStatus_H3 := "M256_Manag_IDB".M256F_IDB[2].tHMR.dHeadStatus;
       "DB_M256F_Scada".tHMR.rHeadUsage_km_H3 := "M256_Manag_IDB".M256F_IDB[2].tHMR.rHeadUsage_km;
       "DB_M256F_Scada".tHMR.tManCmd.xMan_FireON_Fdbk_H3 := "M256_Manag_IDB".M256F_IDB[2].tHMR.tManCmd.xMan_FireON_Fdbk;
       "DB_M256F_Scada".tHMR.tManCmd.xMan_FireOFF_Fdbk_H3 := "M256_Manag_IDB".M256F_IDB[2].tHMR.tManCmd.xMan_FireOFF_Fdbk;
       "DB_M256F_Scada".tHMR.tManCmd.xMan_OilON_Fdbk_H3 := "M256_Manag_IDB".M256F_IDB[2].tHMR.tManCmd.xMan_OilON_Fdbk;
       //H4
       "DB_M256F_Scada".tHMR.dHeadStatus_H4 := "M256_Manag_IDB".M256F_IDB[3].tHMR.dHeadStatus;
       "DB_M256F_Scada".tHMR.rHeadUsage_km_H4 := "M256_Manag_IDB".M256F_IDB[3].tHMR.rHeadUsage_km;
       "DB_M256F_Scada".tHMR.tManCmd.xMan_FireON_Fdbk_H4 := "M256_Manag_IDB".M256F_IDB[3].tHMR.tManCmd.xMan_FireON_Fdbk;
       "DB_M256F_Scada".tHMR.tManCmd.xMan_FireOFF_Fdbk_H4 := "M256_Manag_IDB".M256F_IDB[3].tHMR.tManCmd.xMan_FireOFF_Fdbk;
       "DB_M256F_Scada".tHMR.tManCmd.xMan_OilON_Fdbk_H4 := "M256_Manag_IDB".M256F_IDB[3].tHMR.tManCmd.xMan_OilON_Fdbk;
       //H5
       "DB_M256F_Scada".tHMR.dHeadStatus_H5 := "M256_Manag_IDB".M256F_IDB[4].tHMR.dHeadStatus;
       "DB_M256F_Scada".tHMR.rHeadUsage_km_H5 := "M256_Manag_IDB".M256F_IDB[4].tHMR.rHeadUsage_km;
       "DB_M256F_Scada".tHMR.tManCmd.xMan_FireON_Fdbk_H5 := "M256_Manag_IDB".M256F_IDB[4].tHMR.tManCmd.xMan_FireON_Fdbk;
       "DB_M256F_Scada".tHMR.tManCmd.xMan_FireOFF_Fdbk_H5 := "M256_Manag_IDB".M256F_IDB[4].tHMR.tManCmd.xMan_FireOFF_Fdbk;
       "DB_M256F_Scada".tHMR.tManCmd.xMan_OilON_Fdbk_H5 := "M256_Manag_IDB".M256F_IDB[4].tHMR.tManCmd.xMan_OilON_Fdbk;
       //H6
       "DB_M256F_Scada".tHMR.dHeadStatus_H6 := "M256_Manag_IDB".M256F_IDB[5].tHMR.dHeadStatus;
       "DB_M256F_Scada".tHMR.rHeadUsage_km_H6 := "M256_Manag_IDB".M256F_IDB[5].tHMR.rHeadUsage_km;
       "DB_M256F_Scada".tHMR.tManCmd.xMan_FireON_Fdbk_H6 := "M256_Manag_IDB".M256F_IDB[5].tHMR.tManCmd.xMan_FireON_Fdbk;
       "DB_M256F_Scada".tHMR.tManCmd.xMan_FireOFF_Fdbk_H6 := "M256_Manag_IDB".M256F_IDB[5].tHMR.tManCmd.xMan_FireOFF_Fdbk;
       "DB_M256F_Scada".tHMR.tManCmd.xMan_OilON_Fdbk_H6 := "M256_Manag_IDB".M256F_IDB[5].tHMR.tManCmd.xMan_OilON_Fdbk;
       //H7
       "DB_M256F_Scada".tHMR.dHeadStatus_H7 := "M256_Manag_IDB".M256F_IDB[6].tHMR.dHeadStatus;
       "DB_M256F_Scada".tHMR.rHeadUsage_km_H7 := "M256_Manag_IDB".M256F_IDB[6].tHMR.rHeadUsage_km;
       "DB_M256F_Scada".tHMR.tManCmd.xMan_FireON_Fdbk_H7 := "M256_Manag_IDB".M256F_IDB[6].tHMR.tManCmd.xMan_FireON_Fdbk;
       "DB_M256F_Scada".tHMR.tManCmd.xMan_FireOFF_Fdbk_H7 := "M256_Manag_IDB".M256F_IDB[6].tHMR.tManCmd.xMan_FireOFF_Fdbk;
       "DB_M256F_Scada".tHMR.tManCmd.xMan_OilON_Fdbk_H7 := "M256_Manag_IDB".M256F_IDB[6].tHMR.tManCmd.xMan_OilON_Fdbk;
       //H8
       "DB_M256F_Scada".tHMR.dHeadStatus_H8 := "M256_Manag_IDB".M256F_IDB[7].tHMR.dHeadStatus;
       "DB_M256F_Scada".tHMR.rHeadUsage_km_H8 := "M256_Manag_IDB".M256F_IDB[7].tHMR.rHeadUsage_km;
       "DB_M256F_Scada".tHMR.tManCmd.xMan_FireON_Fdbk_H8 := "M256_Manag_IDB".M256F_IDB[7].tHMR.tManCmd.xMan_FireON_Fdbk;
       "DB_M256F_Scada".tHMR.tManCmd.xMan_FireOFF_Fdbk_H8 := "M256_Manag_IDB".M256F_IDB[7].tHMR.tManCmd.xMan_FireOFF_Fdbk;
       "DB_M256F_Scada".tHMR.tManCmd.xMan_OilON_Fdbk_H8 := "M256_Manag_IDB".M256F_IDB[7].tHMR.tManCmd.xMan_OilON_Fdbk;




